// TIA Portal project "EbAndon v2_1_0" (V15) (continued)
TYPE "KP8 Button Config"
   STRUCT
      activate : Array[0.."ptsPerStn"] of Bool;
      colorOn1 : Array[0.."ptsPerStn"] of String[10];
      colorOn2 : Array[0.."ptsPerStn"] of String[10];
      colorOff : Array[0.."ptsPerStn"] of String[10];
      flash : Array[0.."ptsPerStn"] of Bool;
      group : Array[0.."ptsPerStn"] of Int;
      mode : Array[0.."ptsPerStn"] of Bool;
   END_STRUCT;
END_TYPE

TYPE "Elapsed Time"
   STRUCT
      partReq : Array[0.."ptsPerStn"] of Real;
      resetReq : Real;
   END_STRUCT;
END_TYPE

TYPE "Part Request Data"
   STRUCT
      row : Array[0.."partReqDataRowCount"] of "Table Row";
   END_STRUCT;
END_TYPE

TYPE "Station"
   STRUCT
      animations : Array[0.."ptsPerStn"] of Int;
      btnStates : Array[0.."ptsPerStn"] of Bool;
      dropZone : USInt;
      elapsedTime : "Elapsed Time";
      groupSelect : Int;
      kp8Config : "KP8 Button Config";
      kp8In : Byte;
      kp8Out : DWord;
      init : "Station Initialization";
      line : WString[20];
      partNumbers : Array[0.."ptsPerStn"] of WString["mStringLen"];
      partOrdered : Array[0.."ptsPerStn"] of Bool;
      partRequested : Array[0.."ptsPerStn"] of Bool;
      presetTime : "Preset Time";
      settings : "Station Settings Screen";
      stackLightOut : DWord;
   END_STRUCT;
END_TYPE

TYPE "Settings"
   STRUCT
      alotted : Struct
         assign : "PB Data: Text Label";
         ioField : "IO Field Data: Timers";
      END_STRUCT;
      critical : Struct
         assign : "PB Data: Text Label";
         ioField : "IO Field Data: Timers";
      END_STRUCT;
      kp8 : Struct
         selectButtons : "PB Data: Text Label";
         btnSelState : Array[0.."ptsPerStn"] of Bool;
         buttons : Array[0.."ptsPerStn"] of "PB Data: Text Label";
         selBtnNumber : Int;
         selCount : Int;
      END_STRUCT;
      stations : Struct
         selectAll : "PB Data: Text Label";
         nextGroup : "PB Data: Graphic/Text List";
         prevGroup : "PB Data: Graphic/Text List";
         selectBtns : Array[0.."hmiSelStnCount"] of "PB Data: Text Label";
         selCount : Int;
         selNumber : Int;
      END_STRUCT;
      partNumber : Struct
         assign : "PB Data: Text Label";
         ioField : "IO Field Data: Part Number";
      END_STRUCT;
      viewingStation : Struct
         btns : Array[0.."ptsPerStn"] of "Station Assignment: Button Details";
         dzData : "Drop Zone Data";
         lineData : "Line Label Data";
         next : "PB Data: Graphic/Text List";
         previous : "PB Data: Graphic/Text List";
         "name" : WString[20];
      END_STRUCT;
   END_STRUCT;
END_TYPE

TYPE "PB Data: Graphic/Text List"
   STRUCT
      actuate : Bool;
      animate : USInt;
      listSelect : UInt;
   END_STRUCT;
END_TYPE

TYPE "LED Sign Data"
   STRUCT
      row : Array[0.."ledRowCount"] of "Table Row";
   END_STRUCT;
END_TYPE

TYPE "PB Data: Text Label"
   STRUCT
      actuate : Bool;
      animate : USInt;
      label : WString[20];
   END_STRUCT;
END_TYPE

TYPE "Station Old Presses"
   STRUCT
      me : Array[0.."stnCount", 0.."ptsPerStn"] of Bool;
   END_STRUCT;
END_TYPE

TYPE "Station Assignment: Button Details"
   STRUCT
      alloted : Struct
         animate : USInt;
         value : WString[10];
      END_STRUCT;
      critical : Struct
         animate : USInt;
         value : WString[10];
      END_STRUCT;
      label : Struct
         animate : USInt;
         value : WString[2];
      END_STRUCT;
      partNumber : Struct
         animate : USInt;
         value : WString[40];
      END_STRUCT;
      select : Struct
         actuate : Bool;
         animate : USInt;
      END_STRUCT;
   END_STRUCT;
END_TYPE

TYPE "IO Field Data: Part Number"
   STRUCT
      animate : USInt;
      inputFinished : Bool;
      value : WString[40];
   END_STRUCT;
END_TYPE

TYPE "Line Label Data"
   STRUCT
      animate : Struct
         bg : USInt;
         ioField : USInt;
      END_STRUCT;
      inputFinished : Bool;
      value : WString[10];
   END_STRUCT;
END_TYPE

TYPE "Drop Zone Data"
   STRUCT
      animate : Struct
         bg : USInt;
         ioField : USInt;
      END_STRUCT;
      inputFinished : Bool;
      value : WString[10];
   END_STRUCT;
END_TYPE

TYPE "IO Field Data: Timers"
   STRUCT
      animate : USInt;
      inputFinished : Bool;
      value : WString[5];
   END_STRUCT;
END_TYPE

TYPE "Table Nav"
   STRUCT
      top : "PB Data: Graphic/Text List";
      pageUp : "PB Data: Graphic/Text List";
      lineUp : "PB Data: Graphic/Text List";
      lineDown : "PB Data: Graphic/Text List";
      pageDown : "PB Data: Graphic/Text List";
      bottom : "PB Data: Graphic/Text List";
   END_STRUCT;
END_TYPE

TYPE "Station Sim Data"
   STRUCT
      stn : Struct
         animate : USInt;
         label : WString[20];
      END_STRUCT;
      btn : Struct
         actuate : Byte;
         animate : Array[0..7] of USInt;
         labels : Array[0..7] of WString [4];
      END_STRUCT;
   END_STRUCT;
END_TYPE

TYPE "Simulated Stations"
   STRUCT
      down : "PB Data: Graphic/Text List";
      firstStn : Int;
      me : Array[0.."simKP8Count"] of "Station Sim Data";
      up : "PB Data: Graphic/Text List";
   END_STRUCT;
END_TYPE

TYPE "Part Req Log"
   STRUCT
      me : Array[0..99] of "Part Req Log Row";
   END_STRUCT;
END_TYPE

TYPE "UserDiag_typeSlot"
   STRUCT
      hardwareId : Hw_Io := 16#0000;   // Hardware identifier of the module which is inserted in the slot
      state : USInt := 0;   // Status of the device/slave. 1:ok; 2:faulty, 3:lost connection, 4:disabled, 5:problem, 12:was faulty, 13:was lost, 14:was disabled, 15:problem gone
      exists : Bool := FALSE;   // TRUE: Modul is existing
      configured : Bool := FALSE;   // TRUE: Modul is configured
      faulty : Bool := FALSE;   // TRUE: Modul is faulty
      problem : Bool := FALSE;   // TRUE: Modul has a problem
      disabled : Bool := FALSE;   // TRUE: Modul is disabled
      error : Bool := FALSE;   // TRUE: Error in module which is inserted in the slot
   END_STRUCT;
END_TYPE

TYPE "UserDiag_typePLC"
   STRUCT
      hardwareId : Hw_Device := 16#0000;   // Hardware identifier of the PLC
      error : Bool := FALSE;   // TRUE: Error in PLC
      actualConfiguredSlots : Int := 0;   // Number of configured local slots at PLC
      slots : Array[0.."USERDIAG_SLOTS_PER_PLC_UPPER_LIM"] of "UserDiag_typeSlot";   // Information of the PLC slots; index = slotnumber; PLC always at slot 1
   END_STRUCT;
END_TYPE

TYPE "UserDiag_typeDevice"
   STRUCT
      hardwareId : Hw_Device := 16#0000;   // Hardware identifier of the device/slave
      number : UInt := 0;   // Profinet device number/Profibus address of the slave
      "name" : WString[20] := WSTRING#'';   // Name of the device/slave
      ipAddress : IP_V4;   // IP address of the device
      state : USInt := 0;   // Status of the device/slave. 1:ok; 2:faulty, 3:lost connection, 4:disabled, 5:problem, 12:was faulty, 13:was lost, 14:was disabled, 15:problem gone
      exists : Bool := FALSE;   // TRUE: Device/slave is existing
      configured : Bool := FALSE;   // TRUE: Device/slave is configured
      faulty : Bool := FALSE;   // TRUE: Device/slave is faulty
      problem : Bool := FALSE;   // TRUE: Device/slave has a problem
      disabled : Bool := FALSE;   // TRUE: Device/slave is disabled
      error : Bool := FALSE;   // TRUE: Error in device/slave
      nextDevice : Int := 0;   // device number of next device
      actualConfiguredSlots : Int := 0;   // Number of configured slots in the device/slave
      slots : Array[0.."USERDIAG_SLOTS_PER_DEVICE_UPPER_LIM"] of "UserDiag_typeSlot";   // Slot information of a device/slave
   END_STRUCT;
END_TYPE

TYPE "UserDiag_typeIOSystem"
   STRUCT
      hardwareId : Hw_IoSystem := 16#0000;   // Hardware identifier of the IO-System/DP-Mastersystem
      number : UInt := 0;   // IO-System/DP-Mastersystem number
      error : Bool := FALSE;   // TRUE: Error in IO-System/DP-Mastersystem
      firstDevice : Int := 0;   // device number (index) of first device in IO System
      lastDevice : Int := 0;   // device number (index) of last device IO System
      actualConfiguredDevices : Int := 0;   // Number of configured devices/slaves in IO-System/DP-Mastersystem
      devices : Array[1.."USERDIAG_DEVICES_PER_IO_SYSTEM_UPPER_LIM"] of "UserDiag_typeDevice";   // Device/Slave information
   END_STRUCT;
END_TYPE

TYPE "Network Health Screen"
   STRUCT
      et200spPopUp : "Station: ET200SP Comm Debug Data";
      kp8PopUp : "Station: KP8 Comm Debug Data";
      pnioDevices : Array[1.."pnioDeviceCount"] of "PB Data: Text Label";
      selectedDevice : Int;
   END_STRUCT;
   // // pnioDevices[1] : volvo1601kp8
   // // pnioDevices[2] : volvo1601et200sp
   // // pnioDevices[3] : volvo1602kp8
   // // pnioDevices[4] : volvo1602et200sp
   // // pnioDevices[5] : volvo1603kp8
   // // pnioDevices[6] : volvo1603et200sp
   // // pnioDevices[7] : volvo1604kp8
   // // pnioDevices[8] : volvo1604et200sp
   // // pnioDevices[9] : volvo1605kp8
   // // pnioDevices[10] : volvo1605et200sp
   // // pnioDevices[11] : volvo1606kp8
   // // pnioDevices[12] : volvo1606et200sp
   // // pnioDevices[13] : volvo1607kp8
   // // pnioDevices[14] : volvo1607et200sp
   // // pnioDevices[15] : volvo1608kp8
   // // pnioDevices[16] : volvo1608et200sp
   // // pnioDevices[17] : volvo1609kp8
   // // pnioDevices[18] : volvo1609et200sp
   // // pnioDevices[19] : volvo1610kp8
   // // pnioDevices[20] : volvo1610et200sp
   // // pnioDevices[21] : volvo1611kp8
   // // pnioDevices[22] : volvo1611et200sp
   // // pnioDevices[23] : chm01kp8
   // // pnioDevices[24] : chm01et200sp
   // // pnioDevices[25] : chm02kp8
   // // pnioDevices[26] : chm02et200sp
   // // pnioDevices[27] : chm03kp8
   // // pnioDevices[28] : chm03et200sp
   // // pnioDevices[29] : chm04kp8
   // // pnioDevices[30] : chm04et200sp
   // // pnioDevices[31] : chm05kp8
   // // pnioDevices[32] : chm05et200sp
   // // pnioDevices[33] : cd001kp8
   // // pnioDevices[34] : cd001et200sp
   // // pnioDevices[35] : cd002kp8
   // // pnioDevices[36] : cd002et200sp
   // // pnioDevices[37] : cd003kp8
   // // pnioDevices[38] : cd003et200sp
   // // pnioDevices[39] : bfl01kp8
   // // pnioDevices[40] : bfl01et200sp
   // // pnioDevices[41] : bfl02kp8
   // // pnioDevices[42] : bfl02et200sp
   // // pnioDevices[43] : bfl03kp8
   // // pnioDevices[44] : bfl03et200sp
   // // pnioDevices[45] : lgs01kp8
   // // pnioDevices[46] : lgs01et200sp
   // // pnioDevices[47] : lgs02kp8
   // // pnioDevices[48] : lgs02et200sp
END_TYPE

TYPE "UserDiag_typeActIOSystem"
   STRUCT
      actIOSystemNumber : Int := 1;   // Number of actual selected IO-system/DP-Mastersystem
      actIODeviceNumbers : Array[1.."pnioDeviceCount"] of UInt;   // Device numbers/profibus addresses of actual selected IO-System/DP-Mastersystem
      actIODeviceState : Array[1.."pnioDeviceCount"] of USInt;   // State of devices/slaves in actual selected IO-System/DP-Mastersystem
      actDeviceSlotsUsed : Array[0.."USERDIAG_SLOTS_PER_SCREEN_UPPER_LIM"] of Bool;   // Used slots of actual selected device/slave
      actDeviceSlotsState : Array[0.."USERDIAG_SLOTS_PER_SCREEN_UPPER_LIM"] of USInt;   // States of actual selected device/slave
   END_STRUCT;
END_TYPE

TYPE "Station: ET200SP Comm Debug Data"
   STRUCT
      dismissPB : Bool;
      IM : "ET200SP: IM Data";
      DQ01 : "ET200SP: DQ Data";
      DQ02 : "ET200SP: DQ Data";
      DQ03 : "ET200SP: DQ Data";
      profinetName : Struct
         animate : USInt;
         label : WString[20];
      END_STRUCT;
      serverModule : "ET200SP: Server Module Data";
   END_STRUCT;
END_TYPE

TYPE "ET200SP: IM Data"
   STRUCT
      bg : USInt;
      error : USInt;
      lnk01 : USInt;
      lnk02 : USInt;
      maint : USInt;
      pwr : USInt;
      run : USInt;
   END_STRUCT;
END_TYPE

TYPE "ET200SP: DQ Data"
   STRUCT
      bg : USInt;
      bgTem : USInt;
      diag : USInt;
      pwr : USInt;
      x0 : USInt;
      x1 : USInt;
      x2 : USInt;
      x3 : USInt;
      x4 : USInt;
      x5 : USInt;
      x6 : USInt;
      x7 : USInt;
   END_STRUCT;
END_TYPE

TYPE "ET200SP: Server Module Data"
   STRUCT
      bg : USInt;
   END_STRUCT;
END_TYPE

TYPE "Station: KP8 Comm Debug Data"
   STRUCT
      dismissPB : Bool;
      profinetName : Struct
         animate : USInt;
         label : WString[20];
      END_STRUCT;
      stencilBackground : USInt;
      X1P1 : Struct
         transmit : USInt;
         receive : USInt;
      END_STRUCT;
      X1P2 : Struct
         transmit : USInt;
         receive : USInt;
      END_STRUCT;
   END_STRUCT;
END_TYPE

TYPE "Station Initialization"
   STRUCT
      hard : Bool;
      soft : Bool;
   END_STRUCT;
END_TYPE

TYPE "Preset Time"
   STRUCT
      allotted : Array[0.."ptsPerStn"] of Real;
      critical : Array[0.."ptsPerStn"] of Real;
   END_STRUCT;
END_TYPE

TYPE "Station Settings Screen"
   STRUCT
      selected : Bool;
      btnSelection : Array[0.."ptsPerStn"] of Bool;
   END_STRUCT;
END_TYPE

// folder: HMI Selection Station

TYPE "HSS: Part Selection Screen"
   STRUCT
      animate : Array[0.."hmiStnPartSelScrnBtnCnt"] of Int;
      pbs : DWord;
      txt : Array[0.."hmiStnPartSelScrnBtnCnt"] of WString [40];
   END_STRUCT;
END_TYPE

TYPE "HSS: Compressed"
   STRUCT
      scrnSlctPrt : "HSS: Part Selection Screen";
      scrnSlctMn : "HSS: Menu Selection Screen";
      scrnTmplt : "HSS: Template Screen";
   END_STRUCT;
END_TYPE

TYPE "HSS: Menu Selection Screen"
   STRUCT
      animate : Array[0.."hmiStnMenuSelScrnBtnCnt"] of Int;
      pbs : DWord;
      txt : Array[0.."hmiStnMenuSelLblCnt"] of WString ["lStringLen"];
   END_STRUCT;
END_TYPE

TYPE "HSS: Template Screen"
   STRUCT
      animate : Array[0.."hmiStnTmpltBtnCnt"] of Int;
      pb : DWord;
      text : Array[0.."hmiStnTmpltBtnCnt"] of WString ["lStringLen"];
   END_STRUCT;
END_TYPE

// folder: Menu System

TYPE "Menu: Libraries"
   STRUCT
      stations : Array[0.."stnCount"] of "Menu: Library";
   END_STRUCT;
   // stations[24].entry[0] := WSTRING#'16.08.208.101.020A$LSA DOC Sleeved Before Forming';
   // stations[24].entry[1] := WSTRING#'16.08.209.031.000C$LDOC Stuffed Shell Before Forming';
   // stations[24].entry[2] := WSTRING#'16.08.209.091.000D$LSA DPF Stuffed (after Hess)';
   // stations[24].entry[3] := WSTRING#'16.08.209.233.000E$LSCR Stuffed Shell- NGK Before Forming';
   // stations[24].entry[4] := WSTRING#'16.08.209.437.000A$LDOC Stuffed Shell Unformed';
   // stations[24].entry[5] := WSTRING#'16.08.210.031.000B$LStuffed Shell DOC';
   // stations[24].entry[6] := WSTRING#'16.08.210.421.500A$LStuffed Shell DOC- 2013';
   // stations[24].entry[7] := WSTRING#'16.08.210.428.000A$LSA DPF Stuffed (after Hess)';
   // stations[24].entry[8] := WSTRING#'16.08.211.801.400A$LSA DOC Sleeved';
   // stations[24].entry[9] := WSTRING#'16.08.211.801.700B$LDPF Stuffed Shell 1 box longs only';
   // stations[24].entry[10] := WSTRING#'16.08.211.806.400B$LSA DPF Stuffed Shell';
   // stations[24].entry[11] := WSTRING#'16.08.216.801.600A$LSA DOC Sleeved DDC 2016 unformed';
   // stations[24].entry[12] := WSTRING#'16.08.216.806.400A$L DPF Sleeved 2016';
   // stations[24].entry[13] := WSTRING#'16.08.217.408.000A$LSA DPF SLEEVED Hess';
   // stations[24].entry[14] := WSTRING#'16.08.217.421.500A$LSA DOC SLEEVED - 2HH 2016';
   // stations[24].entry[15] := WSTRING#'16.08.217.737.000A$LSA DOC SLEEVED - 2V2 2016 unformed';
   // stations[24].entry[16] := WSTRING#'16.32.307.322.210A$LVolvo - ASSY INLET - SUB 8 Unformed';
   // stations[24].entry[17] := WSTRING#'16.32.307.332.400A$LAssembly DPF Canning 2016';
   // stations[24].entry[18] := WSTRING#'16.32.307.472.210A$LSA DOC Canning w/out End Forming';
   // stations[24].entry[19] := WSTRING#'16.32.407.322.210A$LVOLVO DOC STUFFED SHELL UNFORMED';
   // stations[24].entry[20] := WSTRING#'16.08.208.081.000H$LDPF Stuffed Shell 1 box longs only';
   // stations[24].entry[21] := WSTRING#'16.08.208.621.000G$LSA DPF Stuffed Shell';
   // stations[24].entry[22] := WSTRING#'16.32.407.322.300A$LDPF Stuffed Shell: MD13/MD16';
   // stations[24].entry[23] := WSTRING#'16.32.307.332.300A$LDPF Stuffed Shell MD11';
   // stations[25].entry[0] := WSTRING#'16.08.210.421.500A$LStuffed Shell DOC- 2013';
   // stations[25].entry[1] := WSTRING#'16.08.217.421.500A$LSA DOC SLEEVED - 2HH 2016';
   // stations[25].entry[2] := WSTRING#'16.08.217.737.000A$LSA DOC SLEEVED - 2V2 2016 unformed';
   // stations[25].entry[3] := WSTRING#'16.08.208.031.000F$LSCR Stuffed Shell 1 box longs only';
   // stations[25].entry[4] := WSTRING#'16.08.208.651.000G$LStuffed Shell SCR- NGK';
   // stations[25].entry[5] := WSTRING#'16.08.211.803.400A$LSCR Stuffed Shell High Power';
   // stations[25].entry[6] := WSTRING#'16.08.217.233.000A$LSA SCR SLEEVED before FORMING';
   // stations[25].entry[7] := WSTRING#'16.32.606.411.000A$LStuffed Shell - SCR Horizontal';
   // stations[25].entry[8] := WSTRING#'16.32.606.421.000A$LStuffed Shell - SCR Horizontal Long- UNI';
   // stations[25].entry[9] := WSTRING#'16.32.706.311.000A$LSCR Stuffed Shell MD11/13: Vert Short';
   // stations[25].entry[10] := WSTRING#'16.32.706.311.001A$LSCR Stuffed Shell MD11/13: Vert Short';
   // stations[25].entry[11] := WSTRING#'16.32.706.341.000A$LSA SCR Catalyst Module - MD11_MD13 -';
   // stations[25].entry[12] := WSTRING#'16.32.706.401.000A$LSCR Stuffed Shell MD11/13: Australia';
   // stations[26].entry[0] := WSTRING#'16.18.015.420.000A$LSA DOC CANNING 11.25 x 5in -END FORMED-';
   // stations[26].entry[1] := WSTRING#'16.08.211.806.400B$LSA DPF Stuffed Shell';
   // stations[26].entry[2] := WSTRING#'16.08.216.801.600A$LSA DOC Sleeved DDC 2016 unformed';
   // stations[26].entry[3] := WSTRING#'16.08.216.806.400A$L DPF Sleeved 2016';
   // stations[26].entry[4] := WSTRING#'16.08.216.751.100A$LSA Sleeved SCR 2016';
   // stations[26].entry[5] := WSTRING#'16.18.007.300.000A$LSA SCR CANNING 9.5 x 10in -END FORMED-';
   // stations[26].entry[6] := WSTRING#'16.18.007.310.000A$LSA SCR CANNING 9.5 x 12in -END FORMED-';
   // stations[26].entry[7] := WSTRING#'16.18.007.320.000B$LSA SCR CANNING 9.5 x 9in -END FORMED-';
   // stations[26].entry[8] := WSTRING#'16.18.008.300.000A$LSA SCR CANNING 9.5 x 12in -END FORMED-';
   // stations[26].entry[9] := WSTRING#'16.18.008.310.000A$LSA SCR CANNING 9.5 x 10in -END FORMED-';
   // stations[26].entry[10] := WSTRING#'16.18.008.320.000A$LSA SCR CANNING 9.5 x 13in -END FORMED-';
   // stations[26].entry[11] := WSTRING#'16.18.008.340.000A$LSA SCR CANNING 9.5 x 13in -END FORMED-';
   // stations[26].entry[12] := WSTRING#'16.18.009.301.000H$LSA SCR CANNING 13 x 11in UNFORMED-';
   // stations[26].entry[13] := WSTRING#'16.18.009.311.000H$LSA SCR CANNING 13 x 12in UNFORMED-';
   // stations[26].entry[14] := WSTRING#'16.18.009.321.000G$LSA SCR CANNING 13 x 9in UNFORMED';
   // stations[26].entry[15] := WSTRING#'16.18.009.331.000F$LSA SCR CANNING 13 x 9in UNFORMED';
   // stations[26].entry[16] := WSTRING#'16.18.009.371.000D$LSA SCR CANNING 13 X10  UNFORMED';
   // stations[26].entry[17] := WSTRING#'16.18.011.300.000A$LSA SCR CANNING 9.5 x 13.5in -END FORMED-';
   // stations[26].entry[18] := WSTRING#'16.18.011.310.000A$L SA SCR CANNING 9.5 x 10in -END FORMED-';
   // stations[26].entry[19] := WSTRING#'16.18.011.320.000A$LSA SCR CANNING 9_5 x 13in -END FORMED-';
   // stations[26].entry[20] := WSTRING#'16.18.011.330.000A$LSA SCR CANNING 9.5 x 9in -END FORMED-';
   // stations[26].entry[21] := WSTRING#'16.18.012.400.000A$LSA DOC CANNING 9.5 x 4in -END FORMED_';
   // stations[26].entry[22] := WSTRING#'16.18.012.410.000A$LSA DOC CANNING 9.5 x 3.3in -END FORMED-';
   // stations[26].entry[23] := WSTRING#'16.18.012.420.000A$LSA DOC CANNING 9.5 x 4in -END FORMED-';
   // stations[26].entry[24] := WSTRING#'16.18.012.430.000A$LSA DOC CANNING 9.5 x 3.3in -END FORMED-';
   // stations[26].entry[25] := WSTRING#'16.18.012.440.000A$LSA DOC CANNING 9.5 x 5in -END FORMED-';
   // stations[26].entry[26] := WSTRING#'16.18.013.410.000A$LSA DOC CANNING 9_5 x 4_5in -END FORMED-';
   // stations[26].entry[27] := WSTRING#'16.18.013.420.000A$LSA DOC CANNING 9.5 x 5.5in -END FORMED-';
   // stations[26].entry[28] := WSTRING#'16.18.015.400.000A$LSA DOC CANNING 11.25 x 4in -END FORMED-';
   // stations[26].entry[29] := WSTRING#'16.18.015.410.000A$LSA DOC CANNING 11_25 x 5in -END FORMED-';
   // stations[26].entry[30] := WSTRING#'16.18.015.430.000A$LSA DOC CANNING 11.25 x 3.4in -END FORMED';
   // stations[26].entry[31] := WSTRING#'16.18.015.450.000A$LSA DOC CANNING 11.25 x 5in -END FORMED-';
   // stations[26].entry[32] := WSTRING#'16.18.016.400.000A$LSA DOC CANNING 11.25 x 3.4in -END FORMED';
   // stations[26].entry[33] := WSTRING#'16.18.017.300.000A$LSA SCR CANNING 12 x 10in -END FORMED-';
   // stations[26].entry[34] := WSTRING#'16.18.017.310.000A$LSA SCR CANNING 12 x 9in -END FORMED-';
   // stations[26].entry[35] := WSTRING#'16.18.017.321.000F$LSA SCR CANNING 12x7in UNFORMED-';
   // stations[26].entry[36] := WSTRING#'16.18.018.400.000A$LSA DOC CANNING 11.25 x 6.8in -END FORMED';
   // stations[26].entry[37] := WSTRING#'16.18.018.410.000A$LSA DOC CANNING 11.25 x 5in -END FORMED-';
   // stations[26].entry[38] := WSTRING#'16.18.018.420.000A$LSA DOC CANNING 11.25 x 6.8in -END FORMED';
   // stations[26].entry[39] := WSTRING#'16.18.018.440.000A$LSA DOC CANNING 11.25 x 5in -END FORMED-';
   // stations[26].entry[40] := WSTRING#'16.18.011.340.000A$LSCR CANNING 9.5 x 9in -END FORMED-';
   // stations[27].entry[0] := WSTRING#'16.08.211.801.700B$LDPF Stuffed Shell 1 box longs only';
   // stations[27].entry[1] := WSTRING#'16.32.307.322.210A$LVolvo - ASSY INLET - SUB 8 Unformed';
   // stations[27].entry[2] := WSTRING#'16.32.606.411.000A$LStuffed Shell - SCR Horizontal';
   // stations[27].entry[3] := WSTRING#'16.32.112.311.001A$LSA SCR CANNING UNFORMED';
   // stations[27].entry[4] := WSTRING#'16.32.112.553.300C$LSA SCR CANNING A700 UNFORMED';
   // stations[27].entry[5] := WSTRING#'16.32.112.304.008A$LASSY SCR CANNING FORMED';
   // stations[27].entry[6] := WSTRING#'16.32.112.516.000G$LASSY DPF CANNING A700';
   // stations[27].entry[7] := WSTRING#'16.32.112.543.000E$LASSY DOC CANNING A700';
   // stations[28].entry[0] := WSTRING#'11.52.001.312.000B$LSA JL 2.2L DPF CANNING';
   // stations[28].entry[1] := WSTRING#'11.54.007.309.000D$LSTUFFED SHELL ASSEMBLY USA-U625';
   // stations[28].entry[2] := WSTRING#'11.54.007.309.002D$LSTUFFED SHELL ASSEMBLY USA-U625';
   // stations[28].entry[3] := WSTRING#'11.54.007.309.009D$LSTUFFED SHELL ASSEMBLY USA-U625';
END_TYPE

TYPE "Menu: Library"
   STRUCT
      size : Int;
      entry : Array[0.."menuCntPerStn"] of WString["lStringLen"];
   END_STRUCT;
END_TYPE

// folder: Global Data

DATA_BLOCK "EMP IDB"   // DB1
{ S7_Optimized_Access := 'TRUE' }
VERSION : 0.1
// stored: InstanceOfName EMP
"EMP"
BEGIN
   stations.me[0].line := WSTRING#'VOLVO 16';
   stations.me[1].line := WSTRING#'VOLVO 16';
   stations.me[2].line := WSTRING#'VOLVO 16';
   stations.me[0].dropZone := 1;
   stations.me[1].dropZone := 2;
   stations.me[2].dropZone := 3;
   stations.me[3].dropZone := 4;
   stations.me[3].line := WSTRING#'VOLVO 16';
   stations.me[4].dropZone := 5;
   stations.me[4].line := WSTRING#'VOLVO 16';
   stations.me[5].line := WSTRING#'VOLVO 16';
   stations.me[5].dropZone := 6;
   stations.me[6].dropZone := 7;
   stations.me[6].line := WSTRING#'VOLVO 16';
   stations.me[7].dropZone := 8;
   stations.me[7].line := WSTRING#'VOLVO 16';
   stations.me[8].dropZone := 9;
   stations.me[8].line := WSTRING#'VOLVO 16';
   stations.me[9].dropZone := 10;
   stations.me[9].line := WSTRING#'VOLVO 16';
   stations.me[10].dropZone := 11;
   stations.me[10].line := WSTRING#'VOLVO 16';
   stations.me[11].line := WSTRING#'CHM';
   stations.me[11].dropZone := 1;
   stations.me[12].line := WSTRING#'CHM';
   stations.me[12].dropZone := 2;
   stations.me[13].line := WSTRING#'CHM';
   stations.me[13].dropZone := 3;
   stations.me[14].dropZone := 4;
   stations.me[14].line := WSTRING#'CHM';
   stations.me[15].line := WSTRING#'CHM';
   stations.me[15].dropZone := 5;
   stations.me[16].dropZone := 1;
   stations.me[16].line := WSTRING#'CDO';
   stations.me[17].dropZone := 2;
   stations.me[17].line := WSTRING#'CDO';
   stations.me[18].line := WSTRING#'CDO';
   stations.me[18].dropZone := 3;
   stations.me[19].dropZone := 1;
   stations.me[19].line := WSTRING#'BFL';
   stations.me[20].dropZone := 2;
   stations.me[20].line := WSTRING#'BFL';
   stations.me[21].line := WSTRING#'BFL';
   stations.me[21].dropZone := 3;
   stations.me[22].dropZone := 1;
   stations.me[22].line := WSTRING#'LGS';
   stations.me[23].line := WSTRING#'LGS';
   stations.me[23].dropZone := 2;
END_DATA_BLOCK

DATA_BLOCK "HMI"   // DB2
{ S7_Optimized_Access := 'TRUE' }
VERSION : 0.1
   VAR
      barcode : "Barcode Screen";
      networkHealth : "Network Health Screen";
      partCall : "Part Call Screen";
      screenNumber : Int;
      settings : "Settings";
      simStations : "Simulated Stations";
      tableNav : "Table Nav";
   END_VAR
BEGIN
END_DATA_BLOCK

DATA_BLOCK "Parts"   // DB3
{ S7_Optimized_Access := 'TRUE' }
VERSION : 0.1
   VAR
      pRow : Int;
   END_VAR
   VAR RETAIN
      requests : "Part Request Data";
   END_VAR
BEGIN
END_DATA_BLOCK

DATA_BLOCK "LED Sign"   // DB4
{ S7_Optimized_Access := 'TRUE' }
VERSION : 0.1
   VAR
      request : "LED Sign Data";
   END_VAR
BEGIN
END_DATA_BLOCK

DATA_BLOCK "Log Buffer"   // DB5
{ S7_Optimized_Access := 'TRUE' }
VERSION : 0.1
   VAR RETAIN
      logFlag : Int;
      partReq : "Part Req Log";
   END_VAR
BEGIN
END_DATA_BLOCK

DATA_BLOCK "HMI Select Stations"   // DB6
{ S7_Optimized_Access := 'TRUE' }
VERSION : 0.1
   VAR
      me : Array[0.."hmiStnCount"] of "HSS: Compressed";
   END_VAR
BEGIN
END_DATA_BLOCK

DATA_BLOCK "Menu Libraries"   // DB9
{ S7_Optimized_Access := 'TRUE' }
VERSION : 0.1
   VAR
      me : "Menu: Libraries";
   END_VAR
BEGIN
   me.stations[24].entry[0] := WSTRING#'16.08.208.101.020A$L$$SA DOC Sleeved Before Forming';
   me.stations[24].entry[1] := WSTRING#'16.08.209.031.000C$LDOC Stuffed Shell Before Forming';
   me.stations[24].entry[2] := WSTRING#'16.08.209.091.000D$LSA DPF Stuffed (after Hess)';
   me.stations[24].entry[3] := WSTRING#'16.08.209.233.000E$LSCR Stuffed Shell- NGK Before Forming';
   me.stations[24].entry[4] := WSTRING#'16.08.209.437.000A$LDOC Stuffed Shell Unformed';
   me.stations[24].entry[5] := WSTRING#'16.08.210.031.000B$LStuffed Shell DOC';
   me.stations[24].entry[6] := WSTRING#'16.08.210.421.500A$LStuffed Shell DOC- 2013';
   me.stations[24].entry[7] := WSTRING#'16.08.210.428.000A$LSA DPF Stuffed (after Hess)';
   me.stations[24].entry[8] := WSTRING#'16.08.211.801.400A$L$$SA DOC Sleeved';
   me.stations[24].entry[9] := WSTRING#'16.08.211.801.700B$LDPF Stuffed Shell 1 box longs only';
   me.stations[24].entry[10] := WSTRING#'16.08.211.806.400B$L$$SA DPF Stuffed Shell';
   me.stations[24].entry[11] := WSTRING#'16.08.216.801.600A$LSA DOC Sleeved DDC 2016 unformed';
   me.stations[24].entry[12] := WSTRING#'16.08.216.806.400A$L DPF Sleeved 2016';
   me.stations[24].entry[13] := WSTRING#'16.08.217.408.000A$LSA DPF SLEEVED Hess';
   me.stations[24].entry[14] := WSTRING#'16.08.217.421.500A$LSA DOC SLEEVED - 2HH 2016';
   me.stations[24].entry[15] := WSTRING#'16.08.217.737.000A$LSA DOC SLEEVED - 2V2 2016 unformed';
   me.stations[24].entry[16] := WSTRING#'16.32.307.322.210A$LVolvo - ASSY INLET - SUB 8 Unformed';
   me.stations[24].entry[17] := WSTRING#'16.32.307.332.400A$LAssembly DPF Canning 2016';
   me.stations[24].entry[18] := WSTRING#'16.32.307.472.210A$LSA DOC Canning w/out End Forming';
   me.stations[24].entry[19] := WSTRING#'16.32.407.322.210A$LVOLVO DOC STUFFED SHELL UNFORMED';
   me.stations[24].entry[20] := WSTRING#'16.08.208.081.000H$LDPF Stuffed Shell 1 box longs only';
   me.stations[24].entry[21] := WSTRING#'16.08.208.621.000G$LSA DPF Stuffed Shell';
   me.stations[24].entry[22] := WSTRING#'16.32.407.322.300A$LDPF Stuffed Shell: MD13/MD16';
   me.stations[24].entry[23] := WSTRING#'16.32.307.332.300A$LDPF Stuffed Shell MD11';
   me.stations[25].entry[0] := WSTRING#'16.08.210.421.500A$LStuffed Shell DOC- 2013';
   me.stations[25].entry[1] := WSTRING#'16.08.217.421.500A$LSA DOC SLEEVED - 2HH 2016';
   me.stations[25].entry[2] := WSTRING#'16.08.217.737.000A$LSA DOC SLEEVED - 2V2 2016 unformed';
   me.stations[25].entry[3] := WSTRING#'16.08.208.031.000F$LSCR Stuffed Shell 1 box longs only';
   me.stations[25].entry[4] := WSTRING#'16.08.208.651.000G$LStuffed Shell SCR- NGK';
   me.stations[25].entry[5] := WSTRING#'16.08.211.803.400A$LSCR Stuffed Shell High Power';
   me.stations[25].entry[6] := WSTRING#'16.08.217.233.000A$LSA SCR SLEEVED before FORMING';
   me.stations[25].entry[7] := WSTRING#'16.32.606.411.000A$LStuffed Shell - SCR Horizontal';
   me.stations[25].entry[8] := WSTRING#'16.32.606.421.000A$LStuffed Shell - SCR Horizontal Long- UNI';
   me.stations[25].entry[9] := WSTRING#'16.32.706.311.000A$L$$SCR Stuffed Shell MD11/13: Vert Short';
   me.stations[25].entry[10] := WSTRING#'16.32.706.311.001A$L$$SCR Stuffed Shell MD11/13: Vert Short';
   me.stations[25].entry[11] := WSTRING#'16.32.706.341.000A$LSA SCR Catalyst Module - MD11_MD13 -';
   me.stations[25].entry[12] := WSTRING#'16.32.706.401.000A$LSCR Stuffed Shell MD11/13: Australia';
   me.stations[26].entry[0] := WSTRING#'16.18.015.420.000A$LSA DOC CANNING 11.25 x 5in -END FORMED-';
   me.stations[26].entry[1] := WSTRING#'16.08.211.806.400B$L$$SA DPF Stuffed Shell';
   me.stations[26].entry[2] := WSTRING#'16.08.216.801.600A$LSA DOC Sleeved DDC 2016 unformed';
   me.stations[26].entry[3] := WSTRING#'16.08.216.806.400A$L DPF Sleeved 2016';
   me.stations[26].entry[4] := WSTRING#'16.08.216.751.100A$LSA Sleeved SCR 2016';
   me.stations[26].entry[5] := WSTRING#'16.18.007.300.000A$LSA SCR CANNING 9.5 x 10in -END FORMED-';
   me.stations[26].entry[6] := WSTRING#'16.18.007.310.000A$LSA SCR CANNING 9.5 x 12in -END FORMED-';
   me.stations[26].entry[7] := WSTRING#'16.18.007.320.000B$LSA SCR CANNING 9.5 x 9in -END FORMED-';
   me.stations[26].entry[8] := WSTRING#'16.18.008.300.000A$LSA SCR CANNING 9.5 x 12in -END FORMED-';
   me.stations[26].entry[9] := WSTRING#'16.18.008.310.000A$LSA SCR CANNING 9.5 x 10in -END FORMED-';
   me.stations[26].entry[10] := WSTRING#'16.18.008.320.000A$LSA SCR CANNING 9.5 x 13in -END FORMED-';
   me.stations[26].entry[11] := WSTRING#'16.18.008.340.000A$LSA SCR CANNING 9.5 x 13in -END FORMED-';
   me.stations[26].entry[12] := WSTRING#'16.18.009.301.000H$LSA SCR CANNING 13 x 11in UNFORMED-';
   me.stations[26].entry[13] := WSTRING#'16.18.009.311.000H$LSA SCR CANNING 13 x 12in UNFORMED-';
   me.stations[26].entry[14] := WSTRING#'16.18.009.321.000G$LSA SCR CANNING 13 x 9in UNFORMED';
   me.stations[26].entry[15] := WSTRING#'16.18.009.331.000F$LSA SCR CANNING 13 x 9in UNFORMED';
   me.stations[26].entry[16] := WSTRING#'16.18.009.371.000D$LSA SCR CANNING 13 X10  UNFORMED';
   me.stations[26].entry[17] := WSTRING#'16.18.011.300.000A$LSA SCR CANNING 9.5 x 13.5in -END FORMED-';
   me.stations[26].entry[18] := WSTRING#'16.18.011.310.000A$L SA SCR CANNING 9.5 x 10in -END FORMED-';
   me.stations[26].entry[19] := WSTRING#'16.18.011.320.000A$LSA SCR CANNING 9_5 x 13in -END FORMED-';
   me.stations[26].entry[20] := WSTRING#'16.18.011.330.000A$LSA SCR CANNING 9.5 x 9in -END FORMED-';
   me.stations[26].entry[21] := WSTRING#'16.18.012.400.000A$LSA DOC CANNING 9.5 x 4in -END FORMED_';
   me.stations[26].entry[22] := WSTRING#'16.18.012.410.000A$LSA DOC CANNING 9.5 x 3.3in -END FORMED-';
   me.stations[26].entry[23] := WSTRING#'16.18.012.420.000A$LSA DOC CANNING 9.5 x 4in -END FORMED-';
   me.stations[26].entry[24] := WSTRING#'16.18.012.430.000A$LSA DOC CANNING 9.5 x 3.3in -END FORMED-';
   me.stations[26].entry[25] := WSTRING#'16.18.012.440.000A$LSA DOC CANNING 9.5 x 5in -END FORMED-';
   me.stations[26].entry[26] := WSTRING#'16.18.013.410.000A$LSA DOC CANNING 9_5 x 4_5in -END FORMED-';
   me.stations[26].entry[27] := WSTRING#'16.18.013.420.000A$LSA DOC CANNING 9.5 x 5.5in -END FORMED-';
   me.stations[26].entry[28] := WSTRING#'16.18.015.400.000A$LSA DOC CANNING 11.25 x 4in -END FORMED-';
   me.stations[26].entry[29] := WSTRING#'16.18.015.410.000A$LSA DOC CANNING 11_25 x 5in -END FORMED-';
   me.stations[26].entry[30] := WSTRING#'16.18.015.430.000A$LSA DOC CANNING 11.25 x 3.4in -END FORMED';
   me.stations[26].entry[31] := WSTRING#'16.18.015.450.000A$LSA DOC CANNING 11.25 x 5in -END FORMED-';
   me.stations[26].entry[32] := WSTRING#'16.18.016.400.000A$LSA DOC CANNING 11.25 x 3.4in -END FORMED';
   me.stations[26].entry[33] := WSTRING#'16.18.017.300.000A$LSA SCR CANNING 12 x 10in -END FORMED-';
   me.stations[26].entry[34] := WSTRING#'16.18.017.310.000A$LSA SCR CANNING 12 x 9in -END FORMED-';
   me.stations[26].entry[35] := WSTRING#'16.18.017.321.000F$LSA SCR CANNING 12x7in UNFORMED-';
   me.stations[26].entry[36] := WSTRING#'16.18.018.400.000A$LSA DOC CANNING 11.25 x 6.8in -END FORMED';
   me.stations[26].entry[37] := WSTRING#'16.18.018.410.000A$LSA DOC CANNING 11.25 x 5in -END FORMED-';
   me.stations[26].entry[38] := WSTRING#'16.18.018.420.000A$LSA DOC CANNING 11.25 x 6.8in -END FORMED';
   me.stations[26].entry[39] := WSTRING#'16.18.018.440.000A$LSA DOC CANNING 11.25 x 5in -END FORMED-';
   me.stations[26].entry[40] := WSTRING#'16.18.011.340.000A$LSCR CANNING 9.5 x 9in -END FORMED-';
   me.stations[27].entry[0] := WSTRING#'16.08.211.801.700B$LDPF Stuffed Shell 1 box longs only';
   me.stations[27].entry[1] := WSTRING#'16.32.307.322.210A$LVolvo - ASSY INLET - SUB 8 Unformed';
   me.stations[27].entry[2] := WSTRING#'16.32.606.411.000A$LStuffed Shell - SCR Horizontal';
   me.stations[27].entry[3] := WSTRING#'16.32.112.311.001A$LSA SCR CANNING UNFORMED';
   me.stations[27].entry[4] := WSTRING#'16.32.112.553.300C$LSA SCR CANNING A700 UNFORMED';
   me.stations[27].entry[5] := WSTRING#'16.32.112.304.008A$LASSY SCR CANNING FORMED';
   me.stations[27].entry[6] := WSTRING#'16.32.112.516.000G$LASSY DPF CANNING A700';
   me.stations[27].entry[7] := WSTRING#'16.32.112.543.000E$LASSY DOC CANNING A700';
   me.stations[28].entry[0] := WSTRING#'11.52.001.312.000B$LSA JL 2.2L DPF CANNING';
   me.stations[28].entry[1] := WSTRING#'11.54.007.309.000D$LSTUFFED SHELL ASSEMBLY USA-U625';
   me.stations[28].entry[2] := WSTRING#'11.54.007.309.002D$LSTUFFED SHELL ASSEMBLY USA-U625';
   me.stations[28].entry[3] := WSTRING#'11.54.007.309.009D$LSTUFFED SHELL ASSEMBLY USA-U625';
   // me.stations[0] : volvo 16 01
   // me.stations[1] : volvo 16 02
   // me.stations[2] : volvo 16 03
   // me.stations[3] : volvo 16 04
   // me.stations[4] : volvo 16 05
   // me.stations[5] : volvo 16 06
   // me.stations[6] : volvo 16 07
   // me.stations[7] : volvo 16 08
   // me.stations[8] : volvo 16 09
   // me.stations[9] : volvo 16 10
   // me.stations[10] : volvo 16 11
   // me.stations[11] : chm 01
   // me.stations[12] : chm 02
   // me.stations[13] : chm 03
   // me.stations[14] : chm 04
   // me.stations[15] : cdo 01
   // me.stations[16] : cdo 02
   // me.stations[17] : cdo 03
   // me.stations[18] : bfl 01
   // me.stations[19] : bfl 02
   // me.stations[20] : bfl 03
   // me.stations[21] : lgs 01
   // me.stations[22] : lgs 02
   // me.stations[23] : lgs 03
   // me.stations[24] : cv 01
   // me.stations[25] : cv 02
   // me.stations[26] : cv 03
   // me.stations[27] : cv 04
   // me.stations[28] : pc 01